REGION Network 8
   RUNG wire#powerrail
      Contact( %XData6.6 )
      { S7_Templates := "SrcType := Int"; S7_GenerateENO := "TRUE" } Add(in1 := 1, in2 := #InOut_1, out => #InOut_1)
   END_RUNG
   // the same network as SCL:
   IF %XData6.6 THEN #InOut_1 := 1 + #InOut_1; END_IF;
END_REGION

REGION Network 9
   RUNG wire#powerrail
      Contact( %XData6.7 )
      { S7_Templates := "SrcType := Int"; S7_GenerateENO := "TRUE" } Add(in1 := 1, in2 := #InOut_1, out => #InOut_1)
   END_RUNG
   // the same network as SCL:
   IF %XData6.7 THEN #InOut_1 := 1 + #InOut_1; END_IF;
END_REGION
END_FUNCTION_BLOCK

// folder: Bloques Estandar/Boosters

FUNCTION "Booster (MTA)" : Void   // FC25, LAD
{ S7_Optimized_Access := 'FALSE' }
VERSION : 0.1
   VAR_TEMP   // added for the SCL form of the ladder/FBD networks
      _w1 : Bool;
      _s5time1 : S5Time;
      _w2 : Bool;
      _s5time2 : S5Time;
      _w3 : Bool;
   END_VAR
BEGIN

REGION Network 1
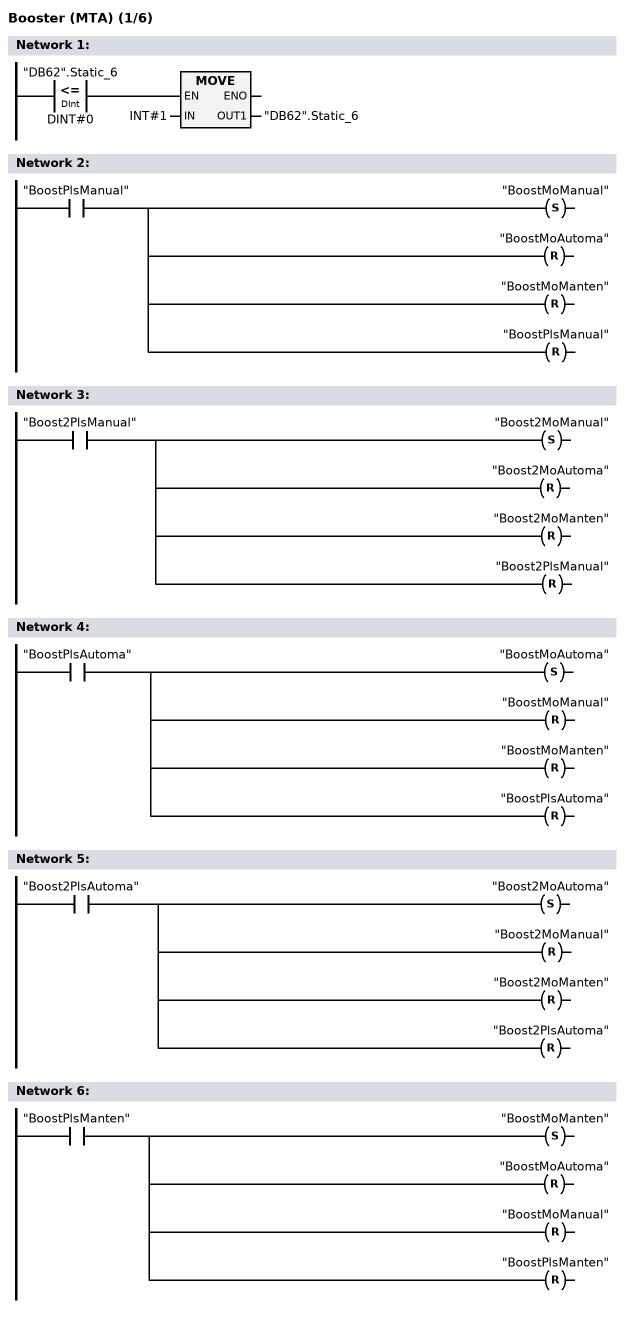
   RUNG wire#powerrail
      { S7_Templates := "SrcType := DInt" } LE_Contact(in1 := "DB62".Static_6, in2 := DINT#0)
      { S7_GenerateENO := "TRUE" } Move(in := INT#1, out1 => "DB62".Static_6)
   END_RUNG
   // the same network as SCL:
   IF "DB62".Static_6 <= DINT#0 THEN "DB62".Static_6 := INT#1; END_IF;
END_REGION

REGION Network 2
   RUNG wire#powerrail
      Contact( "BoostPlsManual" )
      wire#w1
      S_Coil( "BoostMoManual" )
   END_RUNG
   RUNG wire#w1
      R_Coil( "BoostMoAutoma" )
   END_RUNG
   RUNG wire#w1
      R_Coil( "BoostMoManten" )
   END_RUNG
   RUNG wire#w1
      R_Coil( "BoostPlsManual" )
   END_RUNG
   // the same network as SCL:
   IF "BoostPlsManual" THEN
       "BoostMoManual" := TRUE;
       "BoostMoAutoma" := FALSE;
       "BoostMoManten" := FALSE;
       "BoostPlsManual" := FALSE;
   END_IF;
END_REGION

REGION Network 3
   RUNG wire#powerrail
      Contact( "Boost2PlsManual" )
      wire#w1
      S_Coil( "Boost2MoManual" )
   END_RUNG
   RUNG wire#w1
      R_Coil( "Boost2MoAutoma" )
   END_RUNG
   RUNG wire#w1
      R_Coil( "Boost2MoManten" )
   END_RUNG
   RUNG wire#w1
      R_Coil( "Boost2PlsManual" )
   END_RUNG
   // the same network as SCL:
   IF "Boost2PlsManual" THEN
       "Boost2MoManual" := TRUE;
       "Boost2MoAutoma" := FALSE;
       "Boost2MoManten" := FALSE;
       "Boost2PlsManual" := FALSE;
   END_IF;
END_REGION

REGION Network 4
   RUNG wire#powerrail
      Contact( "BoostPlsAutoma" )
      wire#w1
      S_Coil( "BoostMoAutoma" )
   END_RUNG
   RUNG wire#w1
      R_Coil( "BoostMoManual" )
   END_RUNG
   RUNG wire#w1
      R_Coil( "BoostMoManten" )
   END_RUNG
   RUNG wire#w1
      R_Coil( "BoostPlsAutoma" )
   END_RUNG
   // the same network as SCL:
   IF "BoostPlsAutoma" THEN
       "BoostMoAutoma" := TRUE;
       "BoostMoManual" := FALSE;
       "BoostMoManten" := FALSE;
       "BoostPlsAutoma" := FALSE;
   END_IF;
END_REGION

REGION Network 5
   RUNG wire#powerrail
      Contact( "Boost2PlsAutoma" )
      wire#w1
      S_Coil( "Boost2MoAutoma" )
   END_RUNG
   RUNG wire#w1
      R_Coil( "Boost2MoManual" )
   END_RUNG
   RUNG wire#w1
      R_Coil( "Boost2MoManten" )
   END_RUNG
   RUNG wire#w1
      R_Coil( "Boost2PlsAutoma" )
   END_RUNG
   // the same network as SCL:
   IF "Boost2PlsAutoma" THEN
       "Boost2MoAutoma" := TRUE;
       "Boost2MoManual" := FALSE;
       "Boost2MoManten" := FALSE;
       "Boost2PlsAutoma" := FALSE;
   END_IF;
END_REGION

REGION Network 6
   RUNG wire#powerrail
      Contact( "BoostPlsManten" )
      wire#w1
      S_Coil( "BoostMoManten" )
   END_RUNG
   RUNG wire#w1
      R_Coil( "BoostMoAutoma" )
   END_RUNG
   RUNG wire#w1
      R_Coil( "BoostMoManual" )
   END_RUNG
   RUNG wire#w1
      R_Coil( "BoostPlsManten" )
   END_RUNG
   // the same network as SCL:
   IF "BoostPlsManten" THEN
       "BoostMoManten" := TRUE;
       "BoostMoAutoma" := FALSE;
       "BoostMoManual" := FALSE;
       "BoostPlsManten" := FALSE;
   END_IF;
END_REGION

REGION Network 7
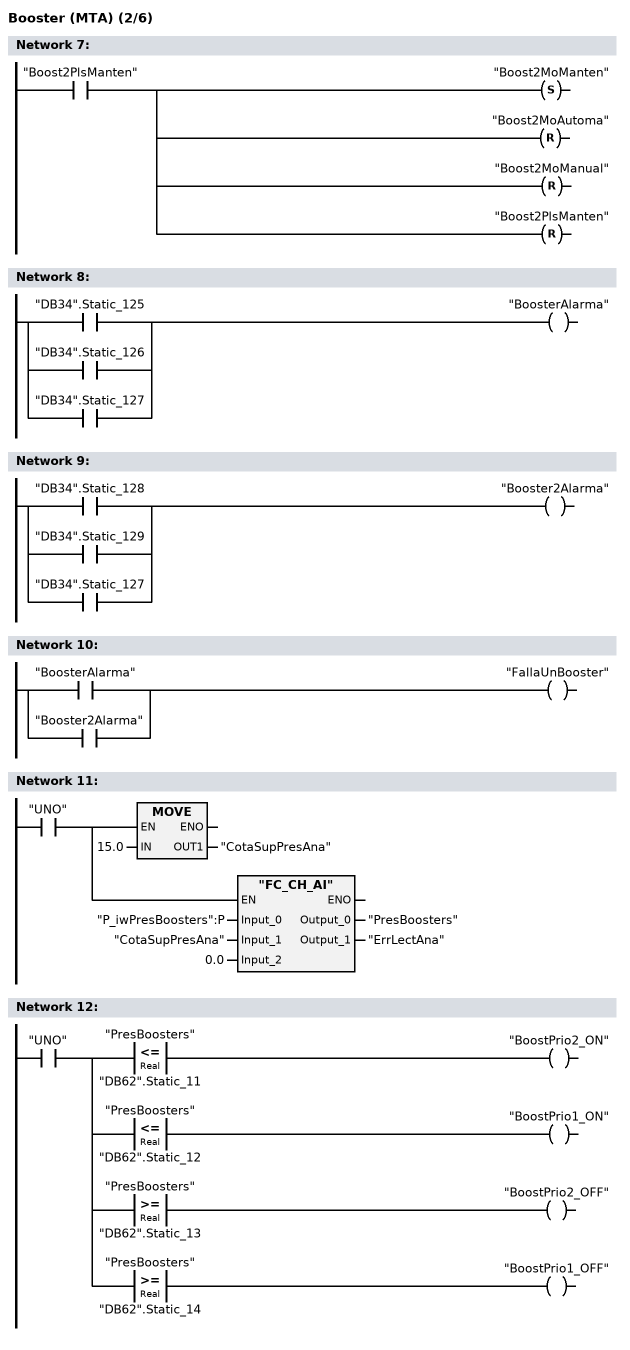
   RUNG wire#powerrail
      Contact( "Boost2PlsManten" )
      wire#w1
      S_Coil( "Boost2MoManten" )
   END_RUNG
   RUNG wire#w1
      R_Coil( "Boost2MoAutoma" )
   END_RUNG
   RUNG wire#w1
      R_Coil( "Boost2MoManual" )
   END_RUNG
   RUNG wire#w1
      R_Coil( "Boost2PlsManten" )
   END_RUNG
   // the same network as SCL:
   IF "Boost2PlsManten" THEN
       "Boost2MoManten" := TRUE;
       "Boost2MoAutoma" := FALSE;
       "Boost2MoManual" := FALSE;
       "Boost2PlsManten" := FALSE;
   END_IF;
END_REGION

REGION Network 8
   RUNG wire#powerrail
      Contact( "DB34".Static_125 )
      wire#w1
      Coil( "BoosterAlarma" )
   END_RUNG
   RUNG wire#powerrail
      Contact( "DB34".Static_126 )
   END_RUNG wire#w1
   RUNG wire#powerrail
      Contact( "DB34".Static_127 )
   END_RUNG wire#w1
   // the same network as SCL:
   "BoosterAlarma" := "DB34".Static_125 OR "DB34".Static_126 OR "DB34".Static_127;
END_REGION

REGION Network 9
   RUNG wire#powerrail
      Contact( "DB34".Static_128 )
      wire#w1
      Coil( "Booster2Alarma" )
   END_RUNG
   RUNG wire#powerrail
      Contact( "DB34".Static_129 )
   END_RUNG wire#w1
   RUNG wire#powerrail
      Contact( "DB34".Static_127 )
   END_RUNG wire#w1
   // the same network as SCL:
   "Booster2Alarma" := "DB34".Static_128 OR "DB34".Static_129 OR "DB34".Static_127;
END_REGION

REGION Network 10
   RUNG wire#powerrail
      Contact( "BoosterAlarma" )
      wire#w1
      Coil( "FallaUnBooster" )
   END_RUNG
   RUNG wire#powerrail
      Contact( "Booster2Alarma" )
   END_RUNG wire#w1
   // the same network as SCL:
   "FallaUnBooster" := "BoosterAlarma" OR "Booster2Alarma";
END_REGION

REGION Network 11
   RUNG wire#powerrail
      Contact( "UNO" )
      wire#w1
      { S7_GenerateENO := "TRUE" } Move(in := 15.0, out1 => "CotaSupPresAna")
   END_RUNG
   RUNG wire#w1
      "FC_CH_AI"(Input_0 := "P_iwPresBoosters":P, Input_1 := "CotaSupPresAna", Input_2 := 0.0, Output_0 => "PresBoosters", Output_1 => "ErrLectAna")
   END_RUNG
   // the same network as SCL:
   IF "UNO" THEN
       "CotaSupPresAna" := 15.0;
       "FC_CH_AI"(Input_0 := "P_iwPresBoosters":P,
                  Input_1 := "CotaSupPresAna",
                  Input_2 := 0.0,
                  Output_0 => "PresBoosters",
                  Output_1 => "ErrLectAna");
   END_IF;
END_REGION

REGION Network 12
   RUNG wire#powerrail
      Contact( "UNO" )
      wire#w1
      { S7_Templates := "SrcType := Real" } LE_Contact(in1 := "PresBoosters", in2 := "DB62".Static_11)
      Coil( "BoostPrio2_ON" )
   END_RUNG
   RUNG wire#w1
      { S7_Templates := "SrcType := Real" } LE_Contact(in1 := "PresBoosters", in2 := "DB62".Static_12)
      Coil( "BoostPrio1_ON" )
   END_RUNG
   RUNG wire#w1
      { S7_Templates := "SrcType := Real" } GE_Contact(in1 := "PresBoosters", in2 := "DB62".Static_13)
      Coil( "BoostPrio2_OFF" )
   END_RUNG
   RUNG wire#w1
      { S7_Templates := "SrcType := Real" } GE_Contact(in1 := "PresBoosters", in2 := "DB62".Static_14)
      Coil( "BoostPrio1_OFF" )
   END_RUNG
   // the same network as SCL:
   "BoostPrio2_ON" := "UNO" AND ("PresBoosters" <= "DB62".Static_11);
   "BoostPrio1_ON" := "UNO" AND ("PresBoosters" <= "DB62".Static_12);
   "BoostPrio2_OFF" := "UNO" AND ("PresBoosters" >= "DB62".Static_13);
   "BoostPrio1_OFF" := "UNO" AND ("PresBoosters" >= "DB62".Static_14);
END_REGION

REGION Network 13
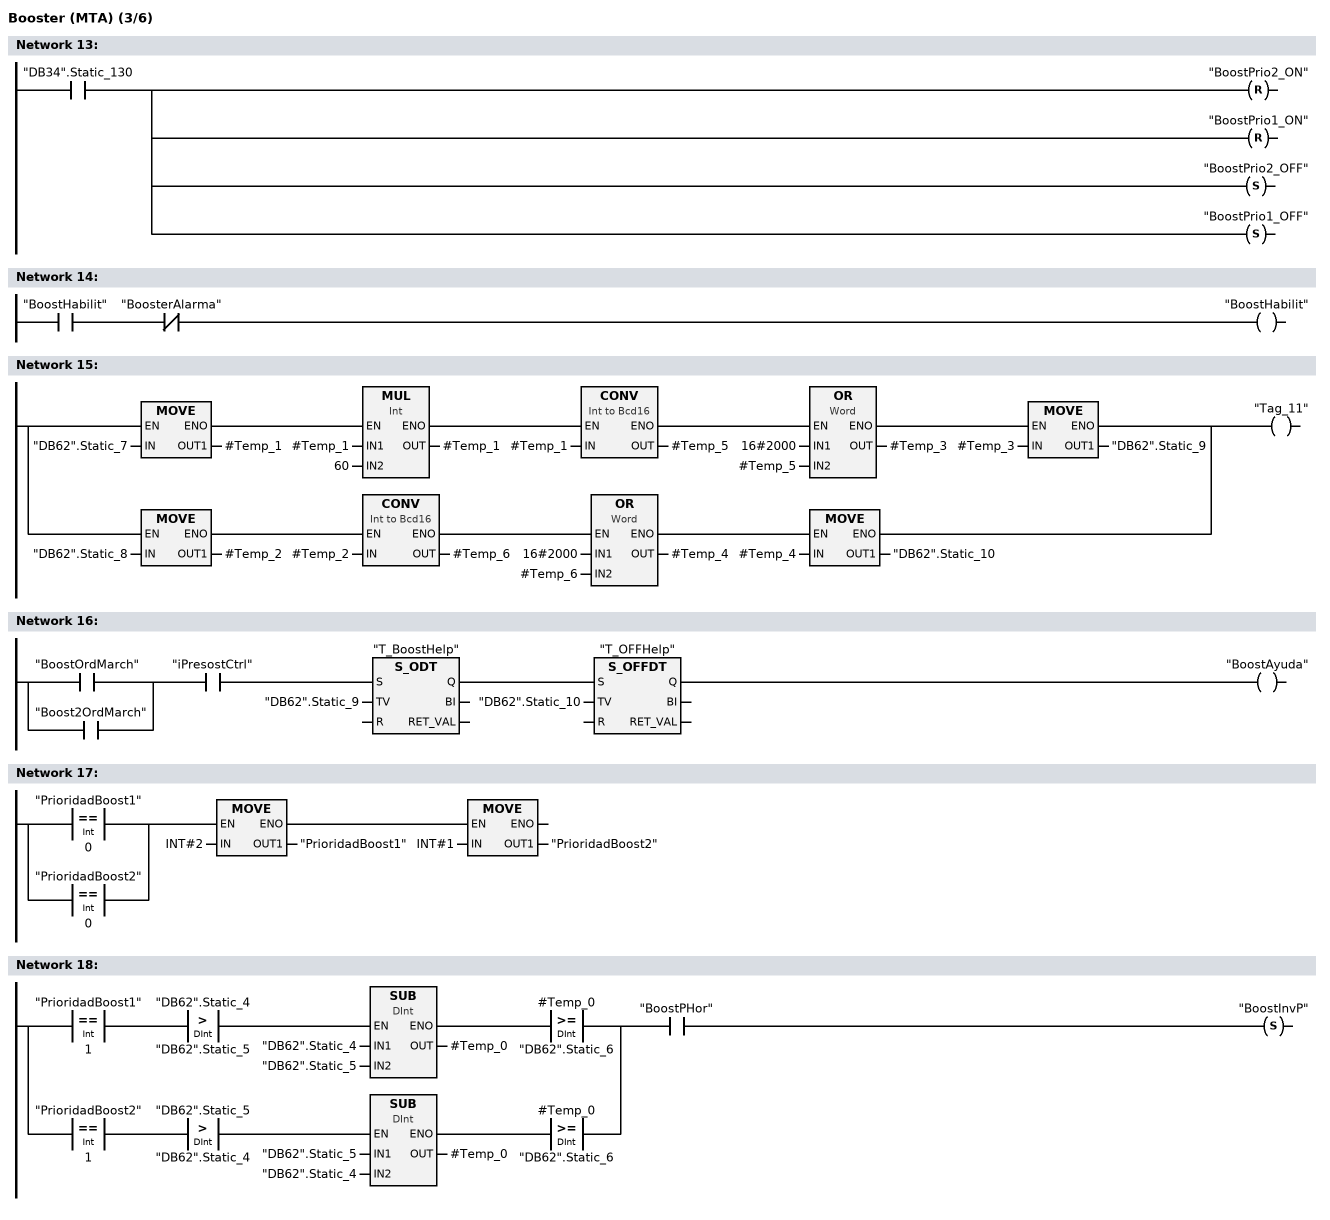
   RUNG wire#powerrail
      Contact( "DB34".Static_130 )
      wire#w1
      R_Coil( "BoostPrio2_ON" )
   END_RUNG
   RUNG wire#w1
      R_Coil( "BoostPrio1_ON" )
   END_RUNG
   RUNG wire#w1
      S_Coil( "BoostPrio2_OFF" )
   END_RUNG
   RUNG wire#w1
      S_Coil( "BoostPrio1_OFF" )
   END_RUNG
   // the same network as SCL:
   IF "DB34".Static_130 THEN
       "BoostPrio2_ON" := FALSE;
       "BoostPrio1_ON" := FALSE;
       "BoostPrio2_OFF" := TRUE;
       "BoostPrio1_OFF" := TRUE;
   END_IF;
END_REGION

REGION Network 14
   RUNG wire#powerrail
      Contact( "BoostHabilit" )
      I_Contact( "BoosterAlarma" )
      Coil( "BoostHabilit" )
   END_RUNG
   // the same network as SCL:
   "BoostHabilit" := "BoostHabilit" AND NOT "BoosterAlarma";
END_REGION

REGION Network 15
   // ENO of a box is taken as its EN; it also drops when the box reports an error
   #Temp_1 := "DB62".Static_7;
   #Temp_1 := #Temp_1 * 60;
   #Temp_5 := INT_TO_BCD16(#Temp_1);
   #Temp_3 := 16#2000 OR #Temp_5;
   "DB62".Static_9 := #Temp_3;
   #Temp_2 := "DB62".Static_8;
   #Temp_6 := INT_TO_BCD16(#Temp_2);
   #Temp_4 := 16#2000 OR #Temp_6;
   "DB62".Static_10 := #Temp_4;
   "Tag_11" := TRUE OR TRUE;
END_REGION

REGION Network 16
   RUNG wire#powerrail
      Contact( "BoostOrdMarch" )
      wire#w1
      Contact( "iPresostCtrl" )
      S_ODT(T_NO := "T_BoostHelp", TV := "DB62".Static_9, R :=, BI =>, RET_VAL =>)
      S_OFFDT(T_NO := "T_OFFHelp", TV := "DB62".Static_10, R :=, BI =>, RET_VAL =>)
      Coil( "BoostAyuda" )
   END_RUNG
   RUNG wire#powerrail
      Contact( "Boost2OrdMarch" )
   END_RUNG wire#w1
   // the same network as SCL:
   #_s5time1 := S_ODT(T_NO := "T_BoostHelp",
                      TV := "DB62".Static_9,
                      S := ("BoostOrdMarch" OR "Boost2OrdMarch") AND "iPresostCtrl",
                      Q => #_w1);
   #_s5time2 := S_OFFDT(T_NO := "T_OFFHelp", S := #_w1, TV := "DB62".Static_10, Q => #_w2);
   "BoostAyuda" := #_w2;
END_REGION

REGION Network 17
   RUNG wire#powerrail
      { S7_Templates := "SrcType := Int" } EQ_Contact(in1 := "PrioridadBoost1", in2 := 0)
      wire#w1
      { S7_GenerateENO := "TRUE" } Move(in := INT#2, out1 => "PrioridadBoost1")
      { S7_GenerateENO := "TRUE" } Move(in := INT#1, out1 => "PrioridadBoost2")
   END_RUNG
   RUNG wire#powerrail
      { S7_Templates := "SrcType := Int" } EQ_Contact(in1 := "PrioridadBoost2", in2 := 0)
   END_RUNG wire#w1
   // the same network as SCL:
   // ENO of a box is taken as its EN; it also drops when the box reports an error
   #_w1 := ("PrioridadBoost1" = 0) OR ("PrioridadBoost2" = 0);
   IF #_w1 THEN
       "PrioridadBoost1" := INT#2;
       "PrioridadBoost2" := INT#1;
   END_IF;
END_REGION

REGION Network 18
   RUNG wire#powerrail
      { S7_Templates := "SrcType := Int" } EQ_Contact(in1 := "PrioridadBoost1", in2 := 1)
      { S7_Templates := "SrcType := DInt" } GT_Contact(in1 := "DB62".Static_4, in2 := "DB62".Static_5)
      { S7_Templates := "SrcType := DInt"; S7_GenerateENO := "TRUE" } Sub(in1 := "DB62".Static_4, in2 := "DB62".Static_5, out => #Temp_0)
      { S7_Templates := "SrcType := DInt" } GE_Contact(in1 := #Temp_0, in2 := "DB62".Static_6)
      wire#w1
      Contact( "BoostPHor" )
      S_Coil( "BoostInvP" )
   END_RUNG
   RUNG wire#powerrail
      { S7_Templates := "SrcType := Int" } EQ_Contact(in1 := "PrioridadBoost2", in2 := 1)
      { S7_Templates := "SrcType := DInt" } GT_Contact(in1 := "DB62".Static_5, in2 := "DB62".Static_4)
      { S7_Templates := "SrcType := DInt"; S7_GenerateENO := "TRUE" } Sub(in1 := "DB62".Static_5, in2 := "DB62".Static_4, out => #Temp_0)
      { S7_Templates := "SrcType := DInt" } GE_Contact(in1 := #Temp_0, in2 := "DB62".Static_6)
   END_RUNG wire#w1
   // the same network as SCL:
   // ENO of a box is taken as its EN; it also drops when the box reports an error
   #_w1 := ("PrioridadBoost1" = 1) AND ("DB62".Static_4 > "DB62".Static_5);
   IF #_w1 THEN #Temp_0 := "DB62".Static_4 - "DB62".Static_5; END_IF;
   #_w2 := ("PrioridadBoost2" = 1) AND ("DB62".Static_5 > "DB62".Static_4);
   #_w3 := #_w1 AND (#Temp_0 >= "DB62".Static_6);
   IF #_w2 THEN #Temp_0 := "DB62".Static_5 - "DB62".Static_4; END_IF;
   IF (#_w3 OR (#_w2 AND (#Temp_0 >= "DB62".Static_6))) AND "BoostPHor" THEN "BoostInvP" := TRUE; END_IF;
END_REGION

REGION Network 19
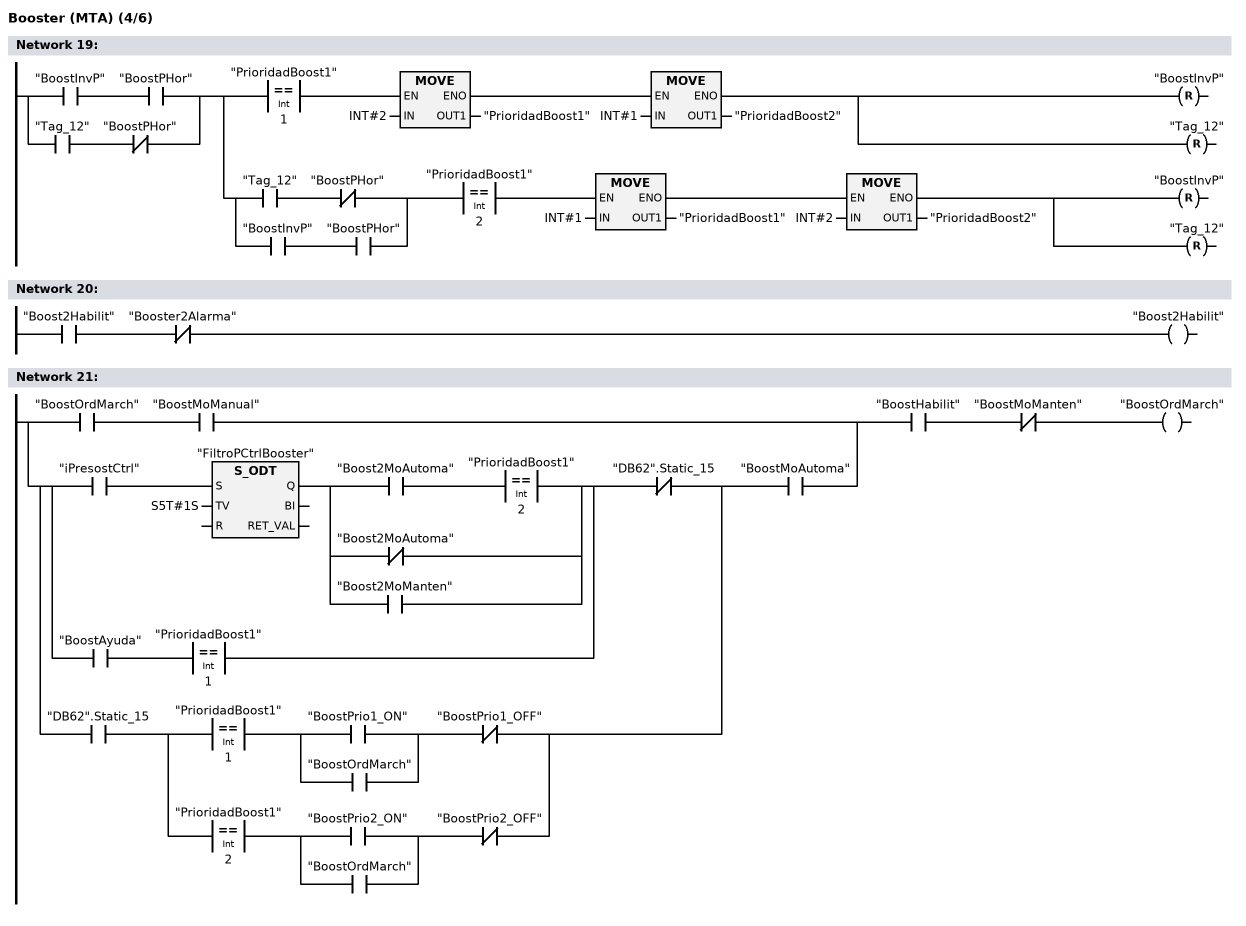
   RUNG wire#powerrail
      Contact( "BoostInvP" )
      Contact( "BoostPHor" )
      wire#w1
      { S7_Templates := "SrcType := Int" } EQ_Contact(in1 := "PrioridadBoost1", in2 := 1)
      { S7_GenerateENO := "TRUE" } Move(in := INT#2, out1 => "PrioridadBoost1")
      { S7_GenerateENO := "TRUE" } Move(in := INT#1, out1 => "PrioridadBoost2")
      wire#w2
      R_Coil( "BoostInvP" )
   END_RUNG
   RUNG wire#powerrail
      Contact( "Tag_12" )
      I_Contact( "BoostPHor" )
   END_RUNG wire#w1
   RUNG wire#w2
      R_Coil( "Tag_12" )
   END_RUNG
   RUNG wire#w1
      Contact( "Tag_12" )
      I_Contact( "BoostPHor" )
      wire#w3
      { S7_Templates := "SrcType := Int" } EQ_Contact(in1 := "PrioridadBoost1", in2 := 2)
      { S7_GenerateENO := "TRUE" } Move(in := INT#1, out1 => "PrioridadBoost1")
      { S7_GenerateENO := "TRUE" } Move(in := INT#2, out1 => "PrioridadBoost2")
      wire#w4
      R_Coil( "BoostInvP" )
   END_RUNG
   RUNG wire#w1
      Contact( "BoostInvP" )
      Contact( "BoostPHor" )
   END_RUNG wire#w3
   RUNG wire#w4
      R_Coil( "Tag_12" )
   END_RUNG
   // the same network as SCL:
   // ENO of a box is taken as its EN; it also drops when the box reports an error
   #_w1 := ("BoostInvP" AND "BoostPHor") OR ("Tag_12" AND NOT "BoostPHor");
   #_w2 := #_w1 AND ("PrioridadBoost1" = 1);
   IF #_w2 THEN
       "PrioridadBoost1" := INT#2;
       "PrioridadBoost2" := INT#1;
       "BoostInvP" := FALSE;
       "Tag_12" := FALSE;
   END_IF;
   #_w3 := #_w1 AND (("Tag_12" AND NOT "BoostPHor") OR ("BoostInvP" AND "BoostPHor")) AND ("PrioridadBoost1" = 2);
   IF #_w3 THEN
       "PrioridadBoost1" := INT#1;
       "PrioridadBoost2" := INT#2;
       "BoostInvP" := FALSE;
       "Tag_12" := FALSE;
   END_IF;
END_REGION

REGION Network 20
   RUNG wire#powerrail
      Contact( "Boost2Habilit" )
      I_Contact( "Booster2Alarma" )
      Coil( "Boost2Habilit" )
   END_RUNG
   // the same network as SCL:
   "Boost2Habilit" := "Boost2Habilit" AND NOT "Booster2Alarma";
END_REGION

REGION Network 21
   #_s5time1 := S_ODT(T_NO := "FiltroPCtrlBooster", TV := S5T#1S, S := "iPresostCtrl", Q => #_w1);
   "BoostOrdMarch" := (("BoostOrdMarch" AND "BoostMoManual") OR (((((#_w1 AND "Boost2MoAutoma" AND ("PrioridadBoost1" = 2)) OR ("BoostAyuda" AND ("PrioridadBoost1" = 1)) OR (#_w1 AND (NOT "Boost2MoAutoma" OR "Boost2MoManten"))) AND NOT "DB62".Static_15) OR ("DB62".Static_15 AND ((("PrioridadBoost1" = 1) AND ("BoostPrio1_ON" OR "BoostOrdMarch") AND NOT "BoostPrio1_OFF") OR (("PrioridadBoost1" = 2) AND ("BoostPrio2_ON" OR "BoostOrdMarch") AND NOT "BoostPrio2_OFF")))) AND "BoostMoAutoma")) AND "BoostHabilit" AND NOT "BoostMoManten";
END_REGION

REGION Network 22
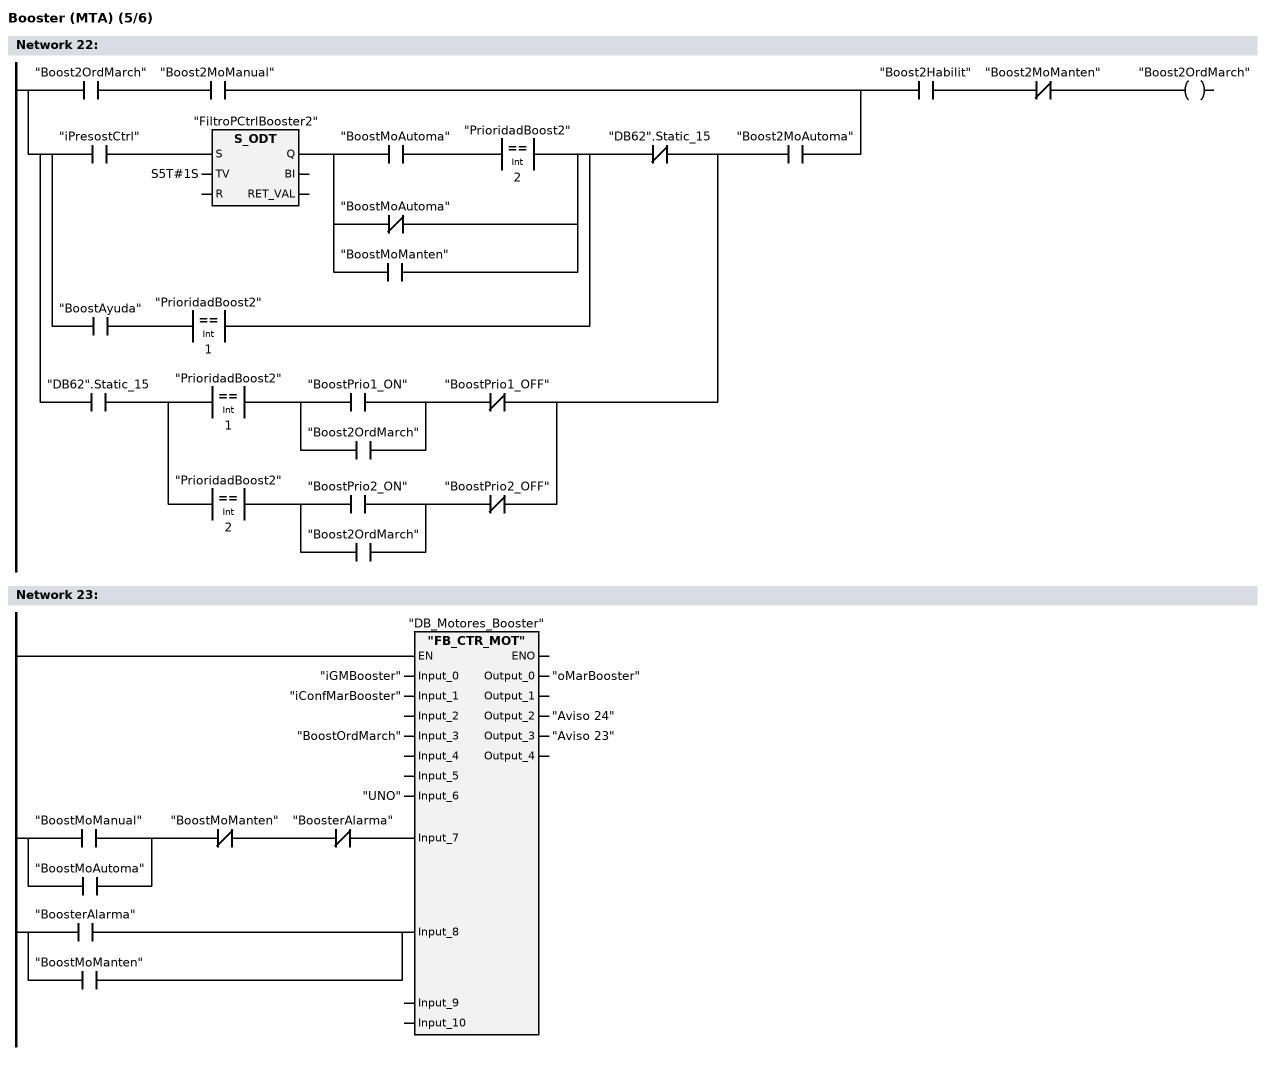
   #_s5time1 := S_ODT(T_NO := "FiltroPCtrlBooster2", TV := S5T#1S, S := "iPresostCtrl", Q => #_w1);
   "Boost2OrdMarch" := (("Boost2OrdMarch" AND "Boost2MoManual") OR (((((#_w1 AND "BoostMoAutoma" AND ("PrioridadBoost2" = 2)) OR ("BoostAyuda" AND ("PrioridadBoost2" = 1)) OR (#_w1 AND (NOT "BoostMoAutoma" OR "BoostMoManten"))) AND NOT "DB62".Static_15) OR ("DB62".Static_15 AND ((("PrioridadBoost2" = 1) AND ("BoostPrio1_ON" OR "Boost2OrdMarch") AND NOT "BoostPrio1_OFF") OR (("PrioridadBoost2" = 2) AND ("BoostPrio2_ON" OR "Boost2OrdMarch") AND NOT "BoostPrio2_OFF")))) AND "Boost2MoAutoma")) AND "Boost2Habilit" AND NOT "Boost2MoManten";
END_REGION

REGION Network 23
   "DB_Motores_Booster"(Input_0 := "iGMBooster",   // "FB_CTR_MOT"
                        Input_1 := "iConfMarBooster",
                        Input_3 := "BoostOrdMarch",
                        Input_6 := "UNO",
                        Input_7 := ("BoostMoManual" OR "BoostMoAutoma") AND NOT "BoostMoManten" AND NOT "BoosterAlarma",
                        Input_8 := "BoosterAlarma" OR "BoostMoManten",
                        Output_0 => "oMarBooster",
                        Output_2 => "Aviso 24",
                        Output_3 => "Aviso 23");
END_REGION

REGION Network 24
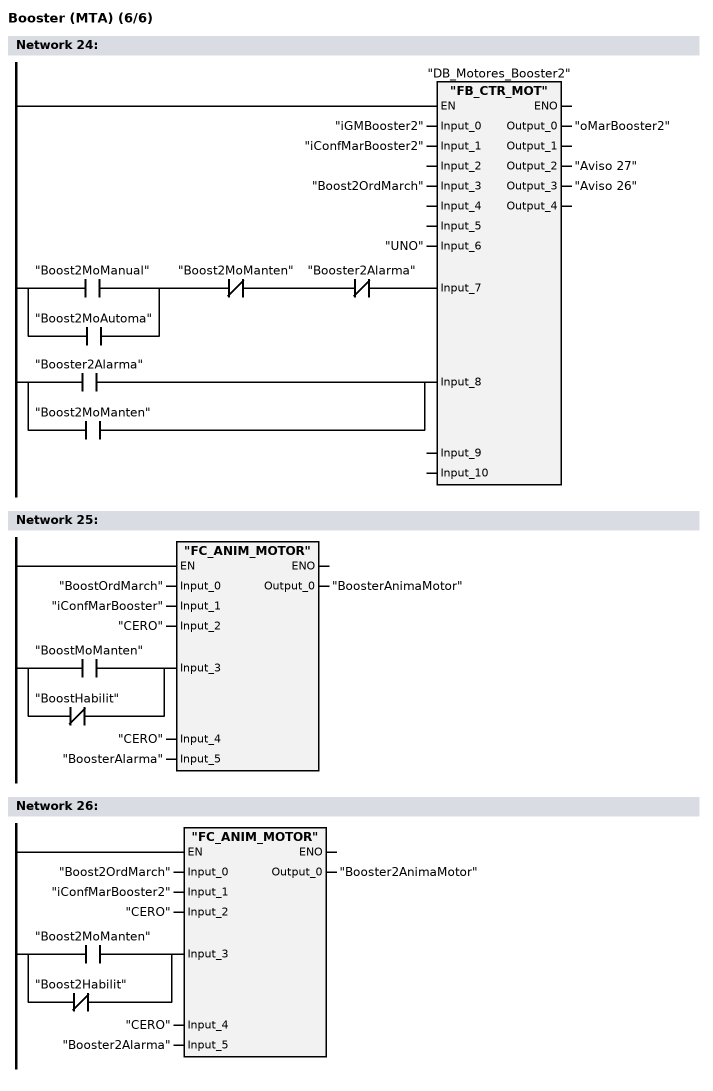
   "DB_Motores_Booster2"(Input_0 := "iGMBooster2",   // "FB_CTR_MOT"
                         Input_1 := "iConfMarBooster2",
                         Input_3 := "Boost2OrdMarch",
                         Input_6 := "UNO",
                         Input_7 := ("Boost2MoManual" OR "Boost2MoAutoma") AND NOT "Boost2MoManten" AND NOT "Booster2Alarma",
                         Input_8 := "Booster2Alarma" OR "Boost2MoManten",
                         Output_0 => "oMarBooster2",
                         Output_2 => "Aviso 27",
                         Output_3 => "Aviso 26");
END_REGION

REGION Network 25
   RUNG wire#powerrail
      "FC_ANIM_MOTOR"(Input_0 := "BoostOrdMarch", Input_1 := "iConfMarBooster", Input_2 := "CERO", Input_3 := wire#w1, Input_4 := "CERO", Input_5 := "BoosterAlarma", Output_0 => "BoosterAnimaMotor")
   END_RUNG
   RUNG wire#powerrail
      Contact( "BoostMoManten" )
   END_RUNG wire#w1
   RUNG wire#powerrail
      I_Contact( "BoostHabilit" )
   END_RUNG wire#w1
   // the same network as SCL:
   "FC_ANIM_MOTOR"(Input_0 := "BoostOrdMarch",
                   Input_1 := "iConfMarBooster",
                   Input_2 := "CERO",
                   Input_3 := "BoostMoManten" OR NOT "BoostHabilit",
                   Input_4 := "CERO",
                   Input_5 := "BoosterAlarma",
                   Output_0 => "BoosterAnimaMotor");
END_REGION

REGION Network 26
   RUNG wire#powerrail
      "FC_ANIM_MOTOR"(Input_0 := "Boost2OrdMarch", Input_1 := "iConfMarBooster2", Input_2 := "CERO", Input_3 := wire#w1, Input_4 := "CERO", Input_5 := "Booster2Alarma", Output_0 => "Booster2AnimaMotor")
   END_RUNG
   RUNG wire#powerrail
      Contact( "Boost2MoManten" )
   END_RUNG wire#w1
   RUNG wire#powerrail
      I_Contact( "Boost2Habilit" )
   END_RUNG wire#w1
   // the same network as SCL:
   "FC_ANIM_MOTOR"(Input_0 := "Boost2OrdMarch",
                   Input_1 := "iConfMarBooster2",
                   Input_2 := "CERO",
                   Input_3 := "Boost2MoManten" OR NOT "Boost2Habilit",
                   Input_4 := "CERO",
                   Input_5 := "Booster2Alarma",
                   Output_0 => "Booster2AnimaMotor");
END_REGION
END_FUNCTION

// folder: Compresores/Alta

FUNCTION "CompresoresAltaMTA" : Void   // FC13, LAD
{ S7_Optimized_Access := 'FALSE' }
VERSION : 0.1
BEGIN

REGION Network 1
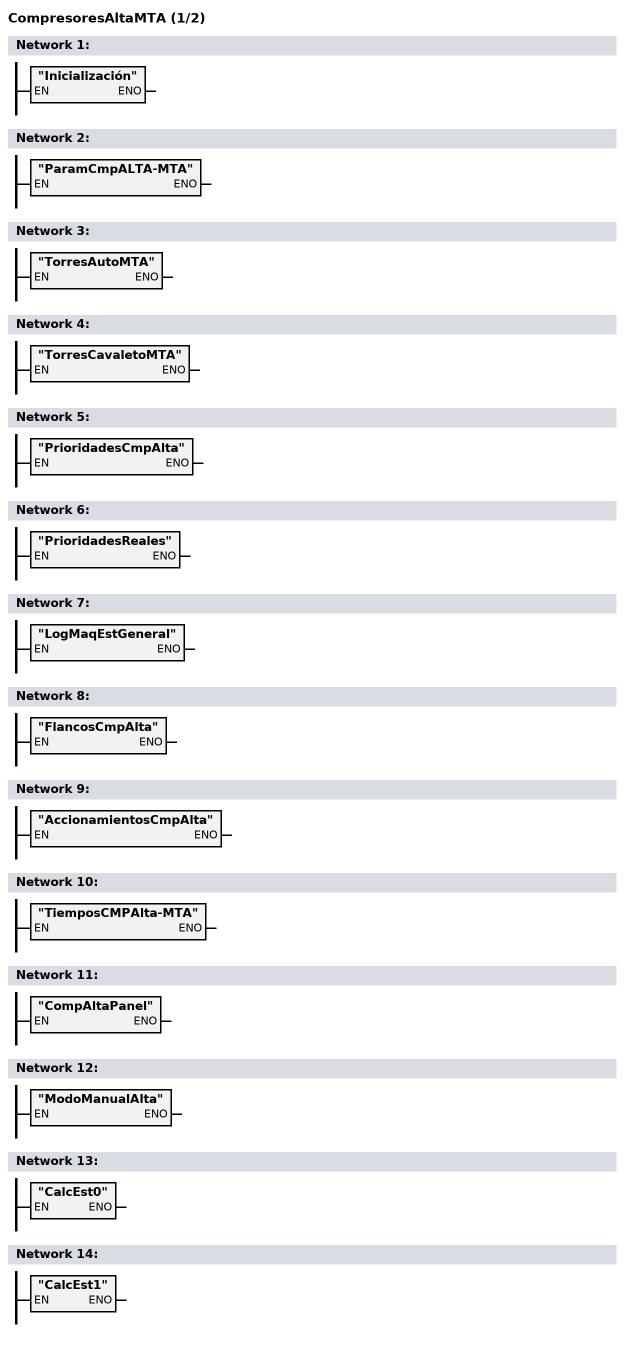
   RUNG wire#powerrail
      "Inicialización"()
   END_RUNG
   // the same network as SCL:
   "Inicialización"();
END_REGION

REGION Network 2
   RUNG wire#powerrail
      "ParamCmpALTA-MTA"()
   END_RUNG
   // the same network as SCL:
   "ParamCmpALTA-MTA"();
END_REGION

REGION Network 3
   RUNG wire#powerrail
      "TorresAutoMTA"()
   END_RUNG
   // the same network as SCL:
   "TorresAutoMTA"();
END_REGION

REGION Network 4
   RUNG wire#powerrail
      "TorresCavaletoMTA"()
   END_RUNG
   // the same network as SCL:
   "TorresCavaletoMTA"();
END_REGION

REGION Network 5
   RUNG wire#powerrail
      "PrioridadesCmpAlta"()
   END_RUNG
   // the same network as SCL:
   "PrioridadesCmpAlta"();
END_REGION

REGION Network 6
   RUNG wire#powerrail
      "PrioridadesReales"()
   END_RUNG
   // the same network as SCL:
   "PrioridadesReales"();
END_REGION

REGION Network 7
   RUNG wire#powerrail
      "LogMaqEstGeneral"()
   END_RUNG
   // the same network as SCL:
   "LogMaqEstGeneral"();
END_REGION

REGION Network 8
   RUNG wire#powerrail
      "FlancosCmpAlta"()
   END_RUNG
   // the same network as SCL:
   "FlancosCmpAlta"();
END_REGION

REGION Network 9
   RUNG wire#powerrail
      "AccionamientosCmpAlta"()
   END_RUNG
   // the same network as SCL:
   "AccionamientosCmpAlta"();
END_REGION

REGION Network 10
   RUNG wire#powerrail
      "TiemposCMPAlta-MTA"()
   END_RUNG
   // the same network as SCL:
   "TiemposCMPAlta-MTA"();
END_REGION

REGION Network 11
   RUNG wire#powerrail
      "CompAltaPanel"()
   END_RUNG
   // the same network as SCL:
   "CompAltaPanel"();
END_REGION

REGION Network 12
   RUNG wire#powerrail
      "ModoManualAlta"()
   END_RUNG
   // the same network as SCL:
   "ModoManualAlta"();
END_REGION

REGION Network 13
   RUNG wire#powerrail
      "CalcEst0"()
   END_RUNG
   // the same network as SCL:
   "CalcEst0"();
END_REGION

REGION Network 14
   RUNG wire#powerrail
      "CalcEst1"()
   END_RUNG
   // the same network as SCL:
   "CalcEst1"();
END_REGION

REGION Network 15
